                 ELSIF #statTokenizedLine.lineToken[#statTokenizedLine.numberOfToken] = #statKeyToken.tokenEndIf
                   AND #statTokenizedLine.numberOfToken = 1
                 THEN
                   REGION ENDIF
                     // EndIF found
                     IF #statStack.numberOfElements > 0 THEN
                       IF #statStack.stackElements[#statStack.numberOfElements].type = "LKINLANG_ENTRY_TYPE_IF" THEN
                         #statStack.stackElements[#statStack.numberOfElements].type := 0;
                         #statStack.stackElements[#statStack.numberOfElements].lineNumberStart := 0;
                         #statStack.numberOfElements -= 1;
                         // go to next state
                         #statStateIntern := #STATE_LINE_PARSED;
                       ELSE
                         // Error not matching stack type 
                         #statStatus := #ERR_PARSING;
                         #statStateIntern := #STATE_ERROR;
                         #statErrorString := CONCAT(IN1 := #statErrorString, IN2 := 'Error: No matching ');
                         #statErrorString := CONCAT(IN1 := #statErrorString, IN2 := #statKeyToken.tokenIf);
                         #statErrorString := CONCAT(IN1 := #statErrorString, IN2 := ' found to ');
                         #statErrorString := CONCAT(IN1 := #statErrorString, IN2 := #statKeyToken.tokenEndIf);
                         #statErrorString := CONCAT(IN1 := #statErrorString, IN2 := ' in line: ');
                         #statErrorString := CONCAT(IN1 := #statErrorString, IN2 := UDINT_TO_STRING(#statTokenizedLine.lineNo));
                       END_IF;
                     ELSE
                       // Error no more elements on stack
                       #statStatus := #ERR_PARSING;
                       #statStateIntern := #STATE_ERROR;
                       #statErrorString := CONCAT(IN1 := #statErrorString, IN2 := 'Error: ');
                       #statErrorString := CONCAT(IN1 := #statErrorString, IN2 := #statKeyToken.tokenEndIf);
                       #statErrorString := CONCAT(IN1 := #statErrorString, IN2 := ' not allowed in line: ');
                       #statErrorString := CONCAT(IN1 := #statErrorString, IN2 := UDINT_TO_STRING(#statTokenizedLine.lineNo));
                     END_IF;
                   END_REGION ENDIF
                 ELSE
                   // Check if line contains WHILE
                   #statStateIntern := #STATE_IS_LINE_WHILE;
                 END_IF;
               END_IF;
             END_REGION IS_LINE_IF

             // ------------------------------------------------------------------------------------------
             // Is line WHILE
             // Check if the line contains WHILE, ENDWHILE
             // If yes then evaluate condition and continue accordingly
             // YES: Go to STATE_LINE_PARSED
             // NO: Go to IS_LINE_FOR
             // ------------------------------------------------------------------------------------------ 
             REGION IS_LINE_WHILE
               IF #statStateIntern = #STATE_IS_LINE_WHILE
               THEN
                 // Definition WHILE:
                 // [1] "10"
                 // [2] ">"
                 // [3] "counter"
                 // [4] " "
                 // [5] "WHILE"
                 // 

                 // Check if line starts with 'WHILE'
                 IF #statTokenizedLine.lineToken[#statTokenizedLine.numberOfToken] = #statKeyToken.tokenWhile THEN
                   REGION WHILE 
                     // WHILE is found
                     // Check if this entry is already on the stack
                     IF #statStack.numberOfElements > 0 THEN
                       IF #statStack.stackElements[#statStack.numberOfElements].lineNumberStart <> #statTokenizedLine.lineNo THEN
                         // New entry on stack
                         #tempReturnVal := 1;
                       ELSE
                         ; // Entry already exists
                       END_IF;
                     ELSE
                       // Empty stack --> Write new entry
                       #tempReturnVal := 1;
                     END_IF;

                     // Create new entry on stack and search matching end
                     IF #tempReturnVal = 1 THEN
                       // Check for ENDWHILE
                       // Search current level of WHILE and find matching ENDWHILE  
                       #tempConditionCounter := -1;
                       FOR #tempCounter := 1 TO #statHierarchicLevel.numberOfLevels DO
                         IF #statHierarchicLevel.levels[#tempCounter].lineNumber = #statTokenizedLine.lineNo THEN
                           #tempConditionCounter := #statHierarchicLevel.levels[#tempCounter].level; // This is the hierarchic level of the current WHILE
                           CONTINUE;
                         END_IF;

                         IF #statHierarchicLevel.levels[#tempCounter].type = "LKINLANG_ENTRY_TYPE_ENDWHILE"
                           AND #statHierarchicLevel.levels[#tempCounter].level = #tempConditionCounter THEN
                           // Correct ENDWHILE found
                           // Exit for loop
                           #tempLineNumber := #statHierarchicLevel.levels[#tempCounter].lineNumber;
                           EXIT;
                         END_IF;
                       END_FOR;

                       // Check if token for ENDWHILE was found
                       IF #tempLineNumber > 0 THEN
                         // New entry on stack
                         #statStack.numberOfElements += 1;
                         IF #statStack.numberOfElements <= "LKINLANG_NUMBER_OF_STACK_ELEMENTS" THEN
                           #statStack.stackElements[#statStack.numberOfElements].type := "LKINLANG_ENTRY_TYPE_WHILE";
                           #statStack.stackElements[#statStack.numberOfElements].lineNumberStart := #statTokenizedLine.lineNo;
                           #statStack.stackElements[#statStack.numberOfElements].lineNumberEnd := #tempLineNumber;
                         ELSE
                           // Error Stack overflow
                           #statStatus := #ERR_PARSING;
                           #statStateIntern := #STATE_ERROR;
                           #statErrorString := CONCAT(IN1 := #statErrorString, IN2 := 'Error: Maximum array index of stack reached');
                           #statErrorString := CONCAT(IN1 := #statErrorString, IN2 := ' in line: ');
                           #statErrorString := CONCAT(IN1 := #statErrorString, IN2 := UDINT_TO_STRING(#statTokenizedLine.lineNo));
                         END_IF;
                       ELSE
                         // Error no ENDWHILE found to WHILE
                         #statStatus := #ERR_PARSING;
                         #statStateIntern := #STATE_ERROR;
                         #statErrorString := CONCAT(IN1 := #statErrorString, IN2 := 'Error: No matching ');
                         #statErrorString := CONCAT(IN1 := #statErrorString, IN2 := #statKeyToken.tokenEndWhile);
                         #statErrorString := CONCAT(IN1 := #statErrorString, IN2 := ' found to ');
                         #statErrorString := CONCAT(IN1 := #statErrorString, IN2 := #statKeyToken.tokenWhile);
                         #statErrorString := CONCAT(IN1 := #statErrorString, IN2 := ' in line: ');
                         #statErrorString := CONCAT(IN1 := #statErrorString, IN2 := UDINT_TO_STRING(#statTokenizedLine.lineNo));
                       END_IF;
                     END_IF;


                     IF #statStateIntern <> #STATE_ERROR THEN
                       // Evaluate the condition and decide where to go next
                       #tempConditionResult := "LKinLang_EvaluateCondition"(offsetLastTokenIndex := 2, // Token offset where condition begins
                                                                            tokenizedLine := #statTokenizedLine,
                                                                            varRefList := #statVarRefList,
                                                                            localVariables := #statVariables,
                                                                            interfaceVariables := #interfaceVariables,
                                                                            keyToken := #statKeyToken,
                                                                            subPrgList := #statSubPrgList,
                                                                            errorString := #statErrorString);

                       // Check if error occured in FC
                       IF #statErrorString <> '' THEN
                         #statStatus := #ERR_PARSING;
                         #statStateIntern := #STATE_ERROR;
                         // Error string was already set
                       END_IF;
                     END_IF;

                     // Check if error was set
                     IF #statStateIntern <> #STATE_ERROR THEN
                       // In case of syntaxCheck being on, always set the condition result to TRUE 
                       // --> Always check if condition
                       IF #statSyntaxCheck <> "LKINLANG_SYNTAX_CHECK_OFF" THEN
                         #tempConditionResult := TRUE;
                       END_IF;

                       // Check the result of the condition
                       IF #tempConditionResult = FALSE THEN
                         // Condition is FALSE --> Go to line after ENDWHILE and remove stack entry
                         #statSearchedLine := #statStack.stackElements[#statStack.numberOfElements].lineNumberEnd + 1;
                         #statStateIntern := #STATE_LINE_PARSED;

                         // Delete stack entry
                         #statStack.stackElements[#statStack.numberOfElements].type := 0;
                         #statStack.stackElements[#statStack.numberOfElements].lineNumberStart := 0;
                         #statStack.stackElements[#statStack.numberOfElements].lineNumberEnd := 0;
                         #statStack.numberOfElements -= 1;
                       ELSE
                         // Condition is TRUE and ENDWHILE is ok --> Nothing more to do
                         #statStateIntern := #STATE_LINE_PARSED;
                       END_IF;
                     END_IF;
                   END_REGION WHILE

                 ELSIF #statTokenizedLine.lineToken[#statTokenizedLine.numberOfToken] = #statKeyToken.tokenEndWhile
                   AND #statTokenizedLine.numberOfToken = 1
                 THEN
                   REGION ENDWHILE
                     // ENDWHILE found --> Can only be found if condition is true 
                     // Check if stack contains correct entry
                     IF #statStack.numberOfElements > 0 THEN
                       IF #statStack.stackElements[#statStack.numberOfElements].type = "LKINLANG_ENTRY_TYPE_WHILE" THEN
                         // Set lineNumber from stack
                         #tempLineNumber := #statStack.stackElements[#statStack.numberOfElements].lineNumberStart;

                         // If syntax check is on then continue in next line
                         IF #statSyntaxCheck = "LKINLANG_SYNTAX_CHECK_OFF" THEN
                           // Go to line containing "WHILE" statement to check condition again
                           #statSearchedLine := #tempLineNumber;
                           #statStateIntern := #STATE_LINE_PARSED;
                         ELSE
                           // Go to next state
                           #statStateIntern := #STATE_LINE_PARSED;
                         END_IF;

                       ELSE
                         // Error not matching stack type 
                         #statStatus := #ERR_PARSING;
                         #statStateIntern := #STATE_ERROR;
                         #statErrorString := CONCAT(IN1 := #statErrorString, IN2 := 'Error: No matching ');
                         #statErrorString := CONCAT(IN1 := #statErrorString, IN2 := #statKeyToken.tokenWhile);
                         #statErrorString := CONCAT(IN1 := #statErrorString, IN2 := ' found to ');
                         #statErrorString := CONCAT(IN1 := #statErrorString, IN2 := #statKeyToken.tokenEndWhile);
                         #statErrorString := CONCAT(IN1 := #statErrorString, IN2 := ' in line: ');
                         #statErrorString := CONCAT(IN1 := #statErrorString, IN2 := UDINT_TO_STRING(#statTokenizedLine.lineNo));
                       END_IF;
                     ELSE
                       // Error no more elements on stack
                       #statStatus := #ERR_PARSING;
                       #statStateIntern := #STATE_ERROR;
                       #statErrorString := CONCAT(IN1 := #statErrorString, IN2 := 'Error: ');
                       #statErrorString := CONCAT(IN1 := #statErrorString, IN2 := #statKeyToken.tokenEndWhile);
                       #statErrorString := CONCAT(IN1 := #statErrorString, IN2 := ' not allowed in line: ');
                       #statErrorString := CONCAT(IN1 := #statErrorString, IN2 := UDINT_TO_STRING(#statTokenizedLine.lineNo));
                     END_IF;
                   END_REGION ENDWHILE
                 ELSE
                   // Parse line token 
                   // Set init state for parsing line token
                   #statStateIntern := #STATE_INIT_PARSE_LOOP;
                   #statStateIntern := #STATE_IS_LINE_FOR;
                 END_IF;
               END_IF;

             END_REGION IS_LINE_WHILE

             // ------------------------------------------------------------------------------------------
             // Is line FOR
             // Check if the line contains FOR, ENDFOR
             // If yes then evaulate FOR loop and continue accordingly
             // YES: Go to STATE_LINE_PARSED
             // NO: Go to IS_LINE_SUB
             // ------------------------------------------------------------------------------------------ 
             REGION IS_LINE_FOR
               IF #statStateIntern = #STATE_IS_LINE_FOR
               THEN
                 // Definition FOR:
                 // SCL: FOR i=10 to 20 by 1 
                 // SIMOTION GCODE: FOR i:10:1:20 // Start:Weite:Ende
                 // FOR i=10,20,1
                 // FOR i:10:20:1

                 // Check if line starts with 'FOR'
                 IF #statTokenizedLine.lineToken[#statTokenizedLine.numberOfToken] = #statKeyToken.tokenFor THEN
                   REGION FOR
                     // FOR is found
                     // Check if this entry is already on the stack
                     IF #statStack.numberOfElements > 0 THEN
                       IF #statStack.stackElements[#statStack.numberOfElements].lineNumberStart <> #statTokenizedLine.lineNo THEN
                         // New entry on stack 
                         #tempReturnVal := 1;
                       ELSE
                         // Entry already exists
                         // Increment counter variable
                         CASE #statStack.stackElements[#statStack.numberOfElements].variableRef.type OF
                           "LKINLANG_VAR_TYPE_LOCAL_DINT":  // Local variable DINT
                             // Local variable at stored index is increased by stored increment
                             #statVariables.dints[#statStack.stackElements[#statStack.numberOfElements].variableRef.index] += #statStack.stackElements[#statStack.numberOfElements].increment;
                           "LKINLANG_VAR_TYPE_INTERFACE_DINT":  // Interface variable DINT
                             // Interface variable at stored index is increased by stored increment
                             #interfaceVariables.DInts[#statStack.stackElements[#statStack.numberOfElements].variableRef.index] += #statStack.stackElements[#statStack.numberOfElements].increment;
                           ELSE  // Wrong variable type
                             ;
                         END_CASE;
                       END_IF;
                     ELSE
                       // Empty stack --> Write new entry
                       #tempReturnVal := 1;
                     END_IF;

                     // -----------------------------------------------------------
                     // New stack entry
                     // -----------------------------------------------------------
                     REGION STACK_ENTRY
                       IF #tempReturnVal = 1 THEN
                         // [1] "1"              --> Step / Increment stored on stack
                         // [2] ":"              --> Delimiter
                         // [3] "20"             --> Target value / Quantitiy stored on stack
                         // [4] ":"              --> Delimiter
                         // [5] "10"             --> Start value
                         // [6] "="              --> Delimiter
                         // [7] "cntr" / "%DI1"  --> Counter variable (must be local or interface(?) variable)
                         // [8] " "
                         // [9] "FOR"

                         // -----------------------------------------------------------
                         // New entry on stack
                         // -----------------------------------------------------------
                         #statStack.numberOfElements += 1;
                         IF #statStack.numberOfElements <= "LKINLANG_NUMBER_OF_STACK_ELEMENTS" THEN
                           #statStack.stackElements[#statStack.numberOfElements].type := "LKINLANG_ENTRY_TYPE_FOR";
                           #statStack.stackElements[#statStack.numberOfElements].lineNumberStart := #statTokenizedLine.lineNo;
                         ELSE
                           // Error Stack overflow
                           #statStatus := #ERR_PARSING;
                           #statStateIntern := #STATE_ERROR;
                           #statErrorString := CONCAT(IN1 := #statErrorString, IN2 := 'Error: Maximum array index of stack reached');
                           #statErrorString := CONCAT(IN1 := #statErrorString, IN2 := ' in line: ');
                           #statErrorString := CONCAT(IN1 := #statErrorString, IN2 := UDINT_TO_STRING(#statTokenizedLine.lineNo));
                           EXIT;
                         END_IF;

                         // -----------------------------------------------------------
                         // SYNTAX: Check correct ENDFOR
                         // -----------------------------------------------------------
                         // Search current level of FOR and find matching ENDFOR
                         #tempConditionCounter := -1;
                         FOR #tempCounter := 1 TO #statHierarchicLevel.numberOfLevels DO
                           IF #statHierarchicLevel.levels[#tempCounter].lineNumber = #statTokenizedLine.lineNo THEN
                             #tempConditionCounter := #statHierarchicLevel.levels[#tempCounter].level; // This is the hierarchic level of the current FOR
                             CONTINUE;
                           END_IF;

                           IF #statHierarchicLevel.levels[#tempCounter].type = "LKINLANG_ENTRY_TYPE_ENDFOR"
                             AND #statHierarchicLevel.levels[#tempCounter].level = #tempConditionCounter THEN
                             // Correct ENDFOR found
                             // Exit for loop
                             #statStack.stackElements[#statStack.numberOfElements].lineNumberEnd := #tempLineNumber := #statHierarchicLevel.levels[#tempCounter].lineNumber;
                             EXIT;
                           END_IF;
                         END_FOR;

                         // Check if token for ENFOR was found
                         IF #tempLineNumber <= 0 THEN
                           // Error no ENDFOR found to FOR
                           #statStatus := #ERR_PARSING;
                           #statStateIntern := #STATE_ERROR;
                           #statErrorString := CONCAT(IN1 := #statErrorString, IN2 := 'Error: No matching ');
                           #statErrorString := CONCAT(IN1 := #statErrorString, IN2 := #statKeyToken.tokenEndFor);
                           #statErrorString := CONCAT(IN1 := #statErrorString, IN2 := ' found to ');
                           #statErrorString := CONCAT(IN1 := #statErrorString, IN2 := #statKeyToken.tokenFor);
                           #statErrorString := CONCAT(IN1 := #statErrorString, IN2 := ' in line: ');
                           #statErrorString := CONCAT(IN1 := #statErrorString, IN2 := UDINT_TO_STRING(#statTokenizedLine.lineNo));
                           EXIT;
                         END_IF;

                         // -----------------------------------------------------------
                         // SYNTAX: Check if space comes after FOR
                         // -----------------------------------------------------------
                         IF #statTokenizedLine.lineToken[#statTokenizedLine.numberOfToken - 1] <> ' ' THEN
                           // Error invalid syntax
                           #statStatus := #ERR_PARSING;
                           #statStateIntern := #STATE_ERROR;
                           #statErrorString := CONCAT(IN1 := #statErrorString, IN2 := 'Error: Invalid syntax in for loop ');
                           #statErrorString := CONCAT(IN1 := #statErrorString, IN2 := ' in line: ');
                           #statErrorString := CONCAT(IN1 := #statErrorString, IN2 := UDINT_TO_STRING(#statTokenizedLine.lineNo));
                           EXIT;
                         END_IF;

                         // -----------------------------------------------------------
                         // SYNTAX: Check if counter can be a variable
                         // -----------------------------------------------------------
                         IF "LKinLang_IsTokenNumberInclSign"(#statTokenizedLine.lineToken[#statTokenizedLine.numberOfToken - 2]) THEN
                           // Error invalid syntax
                           #statStatus := #ERR_PARSING;
                           #statStateIntern := #STATE_ERROR;
                           #statErrorString := CONCAT(IN1 := #statErrorString, IN2 := 'Error: Counter in for loop is not a variable');
                           #statErrorString := CONCAT(IN1 := #statErrorString, IN2 := ' in line: ');
                           #statErrorString := CONCAT(IN1 := #statErrorString, IN2 := UDINT_TO_STRING(#statTokenizedLine.lineNo));
                           EXIT;
                         END_IF;

                         // -----------------------------------------------------------
                         // PARSING: Get counter variable
                         // -----------------------------------------------------------
                         // Copy token to static
                         #statTokenCheck.actual := #statTokenizedLine.lineToken[#statTokenizedLine.numberOfToken - 2];
                         IF #statTokenizedLine.numberOfToken - 3 > 0 THEN
                           #statTokenCheck.previous := #statTokenizedLine.lineToken[#statTokenizedLine.numberOfToken - 3];
                         ELSE
                           #statTokenCheck.previous := '';
                         END_IF;

                         // Check if token is a variable
                         "LKinLang_IsTokenVariable"(lineNumber := #statTokenizedLine.lineNo,
                                                    tokenCheck := #statTokenCheck,
                                                    varIndex => #tempVarIndex,
                                                    varType => #tempVarType,
                                                    varRefList := #statVarRefList,
                                                    keyToken := #statKeyToken,
                                                    subPrgList := #statSubPrgList,
                                                    errorString := #statErrorString,
                                                    stringExpression := #statStringExpression);

                         IF #statErrorString <> '' THEN
                           // Error in function
                           #statStatus := #ERR_PARSING;
                           #statStateIntern := #STATE_ERROR;
                           // String was already set
                           EXIT;
                         ELSIF #tempVarIndex <> 0 AND #tempVarType <> 0 THEN
                           // Variable found
                           // Check if variable is ok --> Store reference on stack
                           IF #tempVarType = "LKINLANG_VAR_TYPE_LOCAL_DINT" OR #tempVarType = "LKINLANG_VAR_TYPE_INTERFACE_DINT" THEN
                             #statStack.stackElements[#statStack.numberOfElements].variableRef.index := #tempVarIndex;
                             #statStack.stackElements[#statStack.numberOfElements].variableRef.type := #tempVarType;
                             //#statStack.stackElements[#statStack.numberOfElements].variableRef.name := ''; // Name is not necessary
                           ELSE
                             // Error: Wrong data type --> Only DINT allowed
                             #statStatus := #ERR_PARSING;
                             #statStateIntern := #STATE_ERROR;
                             #statErrorString := CONCAT(IN1 := #statErrorString, IN2 := 'Error: Invalid data type for counter variable');
                             #statErrorString := CONCAT(IN1 := #statErrorString, IN2 := ' in line: ');
                             #statErrorString := CONCAT(IN1 := #statErrorString, IN2 := UDINT_TO_STRING(#statTokenizedLine.lineNo));
                             EXIT;
                           END_IF;
                         ELSE
                           // Error invalid syntax -> Counter is not a variable
                           #statStatus := #ERR_PARSING;
                           #statStateIntern := #STATE_ERROR;
                           #statErrorString := CONCAT(IN1 := #statErrorString, IN2 := 'Error: Counter in for loop is not a variable');
                           #statErrorString := CONCAT(IN1 := #statErrorString, IN2 := ' in line: ');
                           #statErrorString := CONCAT(IN1 := #statErrorString, IN2 := UDINT_TO_STRING(#statTokenizedLine.lineNo));
                           EXIT;
                         END_IF;

                         // -----------------------------------------------------------
                         // ERROR CHECK: Is counter already used on stack?
                         // -----------------------------------------------------------
                         // Iterate over stack except current entry
                         FOR #tempCounter := 1 TO #statStack.numberOfElements - 1 DO
                           IF #statStack.stackElements[#tempCounter].variableRef.index = #tempVarIndex
                             AND #statStack.stackElements[#tempCounter].variableRef.type = #tempVarType
                           THEN
                             #statStatus := #ERR_PARSING;
                             #statStateIntern := #STATE_ERROR;
                             #statErrorString := CONCAT(IN1 := #statErrorString, IN2 := 'Error: Cannot use same counter in nested for loop');
                             #statErrorString := CONCAT(IN1 := #statErrorString, IN2 := ' in line: ');
                             #statErrorString := CONCAT(IN1 := #statErrorString, IN2 := UDINT_TO_STRING(#statTokenizedLine.lineNo));
                             EXIT;
                           END_IF;
                         END_FOR;

                         IF #statStateIntern = #STATE_ERROR THEN
                           // Abort if error occured
                           EXIT;
                         END_IF;

                         // -----------------------------------------------------------
                         // PARSING: Get delimiters in line
                         // -----------------------------------------------------------
                         // 1:'='
                         // 2:'TO'  // keyToken.tokenQuantity
                         // 3:'STEP'// keyToken.tokenIncrement
                         FOR #tempCounter := #statTokenizedLine.numberOfToken - 3 TO 1 BY -1 DO
                           IF #statTokenizedLine.lineToken[#tempCounter] = '=' AND #tempDelimPos[1] = 0 THEN
                             #tempDelimPos[1] := INT_TO_SINT(#tempCounter);
                           ELSIF #statTokenizedLine.lineToken[#tempCounter] = #statKeyToken.tokenQuantity AND #tempDelimPos[2] = 0 THEN
                             #tempDelimPos[2] := INT_TO_SINT(#tempCounter);
                           ELSIF #statTokenizedLine.lineToken[#tempCounter] = #statKeyToken.tokenIncrement AND #tempDelimPos[3] = 0 THEN
                             #tempDelimPos[3] := INT_TO_SINT(#tempCounter);
                           END_IF;
                         END_FOR;

                         // Check if first delimiter is ok
                         IF #tempDelimPos[1] <= #tempDelimPos[2] OR #tempDelimPos[1] = 0 THEN
                           // ERROR: Wrong delimiter
                           #statStatus := #ERR_PARSING;
                           #statStateIntern := #STATE_ERROR;
                           #statErrorString := CONCAT(IN1 := #statErrorString, IN2 := 'Error: Invalid assignment of start value in for loop');
                           #statErrorString := CONCAT(IN1 := #statErrorString, IN2 := ' in line: ');
                           #statErrorString := CONCAT(IN1 := #statErrorString, IN2 := UDINT_TO_STRING(#statTokenizedLine.lineNo));
                           EXIT;
                         END_IF;

                         // Check if second delimiter is ok
                         IF #tempDelimPos[2] <= #tempDelimPos[3] OR #tempDelimPos[2] = 0 THEN
                           // ERROR: Missing endvalue / quantity
                           #statStatus := #ERR_PARSING;
                           #statStateIntern := #STATE_ERROR;
                           #statErrorString := CONCAT(IN1 := #statErrorString, IN2 := 'Error: Missing quantity in for loop');
                           #statErrorString := CONCAT(IN1 := #statErrorString, IN2 := ' in line: ');
                           #statErrorString := CONCAT(IN1 := #statErrorString, IN2 := UDINT_TO_STRING(#statTokenizedLine.lineNo));
                           EXIT;
                         END_IF;

                         // Check if third delimiter is ok
                         // If not found then increment is set to 1 and parsing increment is skipped 
                         IF #tempDelimPos[3] = 0 THEN
                           #statStack.stackElements[#statStack.numberOfElements].increment := 1; // Inc = 1
                           #tempConditionCounter := 2; // Start with parsing quantity instead of increment
                         ELSE
                           #tempConditionCounter := 3; // Start with parsing increment
                         END_IF;

                         // -----------------------------------------------------------
                         // PARSING: Parse each section between the delimiters
                         // -----------------------------------------------------------
                         #tempTokenCounter := 1; // Init temp
                         // Loop over the necessary variables to parse
                         // 3: Increment (optional)
                         // 2: Quantitiy / EndValue
                         // 1: Start value
                         FOR #tempCounter := #tempConditionCounter TO 1 BY -1 DO

                           // Iterate over all tokens from last delim to next delim
                           WHILE #tempTokenCounter < #tempDelimPos[#tempCounter] DO
                             // Copy token to static
                             #statTokenCheck.actual := #statTokenizedLine.lineToken[#tempTokenCounter];
                             IF #tempTokenCounter > 1 THEN
                               #statTokenCheck.previous := #statTokenizedLine.lineToken[#tempTokenCounter - 1];
                             ELSE
                               #statTokenCheck.previous := '';
                             END_IF;

                             // Skip spaces
                             IF #statTokenCheck.actual = ' ' THEN
                               #tempTokenCounter += 1;
                               CONTINUE;
                             END_IF;

                             // Concat numbers
                             IF "LKinLang_IsTokenNumber"(#statTokenCheck.actual) THEN
                               IF NOT "LKinLang_CharacterIsNumeric"(#statStringExpression[1]) THEN // Check if current stringExpression contains a number
                                 // Not a number --> OK
                                 #statStringExpression := CONCAT(IN1 := #statTokenCheck.actual, IN2 := #statStringExpression);
                                 #tempTokenCounter += 1;
                                 CONTINUE;
                               ELSE
                                 // First char is a number --> Cannot concat two numbers in a row --> ERROR
                                 #statStatus := #ERR_PARSING;
                                 #statStateIntern := #STATE_ERROR;
                                 #statErrorString := CONCAT(IN1 := #statErrorString, IN2 := 'Error: Invalid syntax');
                                 #statErrorString := CONCAT(IN1 := #statErrorString, IN2 := '; Line: ');
                                 #statErrorString := CONCAT(IN1 := #statErrorString, IN2 := UDINT_TO_STRING(#statTokenizedLine.lineNo));
                                 EXIT;
                               END_IF;
                             END_IF;

                             // Check if token is a variable
                             "LKinLang_IsTokenVariable"(lineNumber := #statTokenizedLine.lineNo,
                                                        tokenCheck := #statTokenCheck,
                                                        varIndex => #tempVarIndex,
                                                        varType => #tempVarType,
                                                        varRefList := #statVarRefList,
                                                        keyToken := #statKeyToken,
                                                        subPrgList := #statSubPrgList,
                                                        errorString := #statErrorString,
                                                        stringExpression := #statStringExpression);

                             IF #statErrorString <> '' THEN
                               // Error in function
                               #statStatus := #ERR_PARSING;
                               #statStateIntern := #STATE_ERROR;
                               // String was already set
                               EXIT;
                             ELSIF #tempVarIndex <> 0 AND #tempVarType <> 0 THEN
                               IF NOT "LKinLang_CharacterIsNumeric"(#statStringExpression[1]) THEN
                                 // Variable found --> Get value and concat value to string expression
                                 "LKinLang_GetVariable"(varIndex := #tempVarIndex,
                                                        varType := #tempVarType,
                                                        localVariables := #statVariables,
                                                        interfaceVariables := #interfaceVariables,
                                                        stringExpression := #statStringExpression);
                                 #tempTokenCounter += 1;
                                 CONTINUE;
                               ELSE
                                 // First char is a number --> Cannot concat two numbers in a row --> ERROR
                                 #statStatus := #ERR_PARSING;
                                 #statStateIntern := #STATE_ERROR;
                                 #statErrorString := CONCAT(IN1 := #statErrorString, IN2 := 'Error: Invalid syntax');
                                 #statErrorString := CONCAT(IN1 := #statErrorString, IN2 := '; Line: ');
                                 #statErrorString := CONCAT(IN1 := #statErrorString, IN2 := UDINT_TO_STRING(#statTokenizedLine.lineNo));
                                 EXIT;
                               END_IF;
                             END_IF;

                             // If this section is reached it was not a variable --> Concat
                             // Concat everything else to stringexpression
                             #statStringExpression := CONCAT(IN1 := #statTokenCheck.actual, IN2 := #statStringExpression);
                             #tempTokenCounter += 1;
                             CONTINUE;
                           END_WHILE;

                           // If this section is reached then token counter = delim position
                           // Check if string expression is empty
                           IF #statStringExpression = '' THEN
                             // Error: Empty string!
                             #statStatus := #ERR_PARSING;
                             #statStateIntern := #STATE_ERROR;
                             IF #tempCounter = 1 THEN
                               #statErrorString := CONCAT(IN1 := #statErrorString, IN2 := 'Error: Missing start value assignment in for loop');
                             ELSIF #tempCounter = 2 THEN
                               #statErrorString := CONCAT(IN1 := #statErrorString, IN2 := 'Error: Missing quantity assignment in for loop');
                             ELSE
                               #statErrorString := CONCAT(IN1 := #statErrorString, IN2 := 'Error: Missing increment assignment in for loop');
                             END_IF;
                             #statErrorString := CONCAT(IN1 := #statErrorString, IN2 := ' in line: ');
                             #statErrorString := CONCAT(IN1 := #statErrorString, IN2 := UDINT_TO_STRING(#statTokenizedLine.lineNo));
                             EXIT;
                           END_IF;

                           // Get value of string expression and assign according to counter
                           CASE #tempCounter OF
                             1: // Start value
                               // Assign the start value to the counter variable
                               "LKinLang_SetVariable"(varIndex := #statStack.stackElements[#statStack.numberOfElements].variableRef.index,
                                                      varType := #statStack.stackElements[#statStack.numberOfElements].variableRef.type,
                                                      lineNumber := #statTokenizedLine.lineNo,
                                                      stringExpression := #statStringExpression,
                                                      localVariables := #statVariables,
                                                      interfaceVariables := #interfaceVariables,
                                                      errorString := #statErrorString);

                               IF #statErrorString <> '' THEN // Check if FC has thrown an error
                                 #statStatus := #ERR_PARSING;
                                 #statStateIntern := #STATE_ERROR;
                                 // String was alredy set
                                 EXIT;
                               END_IF;

                             2, 3: // End value & increment
                               // Check if string expression is just a number
                               IF "LKinLang_IsTokenNumberInclSign"(#statStringExpression) THEN
                                 // If just a number then directly assign value
                                 #tempParameterValue := STRING_TO_LREAL(#statStringExpression);
                               ELSE
                                 // Not a single number --> Use mathParser to calculate value
                                 #tempMathParserResult := "LKinLang_CalcMathAndBool"(inputString := #statStringExpression);

                                 // Check for error in math parser
                                 IF #tempMathParserResult.errorID <> 0 THEN
                                   #statErrorString := CONCAT(IN1 := #statErrorString, IN2 := ';Error: Stringexpression ');
                                   #statErrorString := CONCAT(IN1 := #statErrorString, IN2 := #statStringExpression);
                                 ELSE
                                   // Math parser delivers a valid result
                                   // Assign result to value
                                   #tempParameterValue := #tempMathParserResult.finalResult;
                                 END_IF;
                               END_IF;

                               // Check if error occurred
                               IF #statErrorString <> '' THEN
                                 #statStatus := #ERR_PARSING;
                                 #statStateIntern := #STATE_ERROR;
                                 // String was already set
                                 EXIT;
                               ELSE
                                 IF #tempCounter = 2 THEN
                                   // Assign value to quantitiy on stack
                                   #statStack.stackElements[#statStack.numberOfElements].quantity := LREAL_TO_DINT(#tempParameterValue);
                                 ELSE
                                   // Assign value to increment on stack
                                   #statStack.stackElements[#statStack.numberOfElements].increment := LREAL_TO_DINT(#tempParameterValue);
                                   IF #statStack.stackElements[#statStack.numberOfElements].increment = 0 THEN
                                     // ERROR: Increment is 0!
                                     #statStatus := #ERR_PARSING;
                                     #statStateIntern := #STATE_ERROR;
                                     #statErrorString := CONCAT(IN1 := #statErrorString, IN2 := 'Error: Increment in for loop can not be 0');
                                     #statErrorString := CONCAT(IN1 := #statErrorString, IN2 := ' in line: ');
                                     #statErrorString := CONCAT(IN1 := #statErrorString, IN2 := UDINT_TO_STRING(#statTokenizedLine.lineNo));
                                     EXIT;
                                   END_IF;
                                 END_IF;
                               END_IF;
                           END_CASE;

                           // Increment tokenCounter one more time to skip delim
                           #tempTokenCounter += 1;
                           #statStringExpression := '';
                         END_FOR;
                       END_IF;
                     END_REGION STACK_ENTRY


                     // -----------------------------------------------------------
                     // Check the condition -> Counter smaller or equal quantity
                     // YES: Continue in next line (for loop)
                     // NO: Go to endFor (continue after for loop)
                     // -----------------------------------------------------------
                     IF #statStateIntern <> #STATE_ERROR THEN // Check if no error was set
                       // Get value of counter
                       CASE #statStack.stackElements[#statStack.numberOfElements].variableRef.type OF
                         "LKINLANG_VAR_TYPE_LOCAL_DINT":  // Local variable DINT
                           // Get value of local variable
                           #tempParameterValue := #statVariables.dints[#statStack.stackElements[#statStack.numberOfElements].variableRef.index];
                         "LKINLANG_VAR_TYPE_INTERFACE_DINT":  // Interface variable DINT
                           // Get value of interface variable
                           #tempParameterValue := #interfaceVariables.DInts[#statStack.stackElements[#statStack.numberOfElements].variableRef.index];
                         ELSE  // Wrong variable type
                           ;
                       END_CASE;

                       // Check if counting BWD or FWD then check condition accordingly
                       IF #statStack.stackElements[#statStack.numberOfElements].increment > 0 THEN
                         #tempConditionResult := #tempParameterValue <= #statStack.stackElements[#statStack.numberOfElements].quantity;
                       ELSE
                         #tempConditionResult := #tempParameterValue >= #statStack.stackElements[#statStack.numberOfElements].quantity;
                       END_IF;

                       // In case of syntaxCheck being on, always set the condition result to TRUE 
                       // --> Always check if condition
                       IF #statSyntaxCheck <> "LKINLANG_SYNTAX_CHECK_OFF" THEN
                         #tempConditionResult := TRUE;
                       END_IF;

                       // Check the result of the condition
                       IF #tempConditionResult = FALSE THEN
                         // Condition is FALSE --> Go to line after ENDFOR and remove stack entry
                         #statSearchedLine := #statStack.stackElements[#statStack.numberOfElements].lineNumberEnd + 1;
                         #statStateIntern := #STATE_LINE_PARSED;

                         // Delete stack entry
                         #statStack.stackElements[#statStack.numberOfElements].type := 0;
                         #statStack.stackElements[#statStack.numberOfElements].lineNumberStart := 0;
                         #statStack.stackElements[#statStack.numberOfElements].lineNumberEnd := 0;
                         #statStack.stackElements[#statStack.numberOfElements].increment := 0;
                         #statStack.stackElements[#statStack.numberOfElements].quantity := 0;
                         #statStack.stackElements[#statStack.numberOfElements].variableRef.index := 0;
                         #statStack.stackElements[#statStack.numberOfElements].variableRef.type := 0;
                         #statStack.numberOfElements -= 1;

                       ELSE
                         // Condition is TRUE and ENDFOR is ok --> Nothing more to do
                         #statStateIntern := #STATE_LINE_PARSED;
                       END_IF;
                     END_IF;
                   END_REGION FOR

                 ELSIF #statTokenizedLine.lineToken[#statTokenizedLine.numberOfToken] = #statKeyToken.tokenEndFor
                   AND #statTokenizedLine.numberOfToken = 1
                 THEN
                   REGION ENDFOR
                     // ENDFOR found --> ENDFOR is only found if the condition was true, otherwise ENDFOR is skipped 
                     // Check if stack contains correct entry
                     IF #statStack.numberOfElements > 0 THEN
                       IF #statStack.stackElements[#statStack.numberOfElements].type = "LKINLANG_ENTRY_TYPE_FOR" THEN
                         // Set lineNumber from stack but decrease by one as it is increased again outside
                         #tempLineNumber := #statStack.stackElements[#statStack.numberOfElements].lineNumberStart;

                         // If syntax check is on then continue in next line
                         IF #statSyntaxCheck = "LKINLANG_SYNTAX_CHECK_OFF" THEN
                           // Goto line containing the "FOR" statement to check condition again
                           #statSearchedLine := #tempLineNumber;
                           #statStateIntern := #STATE_LINE_PARSED;
                         ELSE
                           // Go to next state
                           #statStateIntern := #STATE_LINE_PARSED;
                         END_IF;